   "Carrier_60_G120DStatusWord.12" AT %I3363.4 : Bool;   // Bit_12_BRAKE_OPEN
   "Carrier_60_G120DStatusWord.13" AT %I3363.5 : Bool;   // Bit_13_NO_OVERTEMP
   "Carrier_60_G120DStatusWord.14" AT %I3363.6 : Bool;   // Bit_14_CW_CCW
   "Carrier_60_G120DStatusWord.15" AT %I3363.7 : Bool;   // Bit_15_OVERL
   "Carrier_60_Slot2_Input" AT %IW3364 : Word;   // SLOT 2 INPUT WORD
   "Carrier_60_CrashDetectSW" AT %I3364.0 : Bool;   // CRASH DETECT SW
   "Carrier_60_SpareSafetyInput(2_1)" AT %I3364.1 : Bool;   // SPARE SAFETY INPUT
   "Carrier_60_SpareSafetyInput(2_2)" AT %I3364.2 : Bool;   // SPARE SAFETY INPUT
   "Carrier_60_SpareSafetyInput(2_3)" AT %I3364.3 : Bool;   // SPARE SAFETY INPUT
   "Carrier_60_SpareSafetyInput(2_4)" AT %I3364.4 : Bool;   // SPARE SAFETY INPUT
   "Carrier_60_SpareSafetyInput(2_5)" AT %I3364.5 : Bool;   // SPARE SAFETY INPUT
   "Carrier_60_SpareSafetyInput(2_6)" AT %I3364.6 : Bool;   // SPARE SAFETY INPUT
   "Carrier_60_SpareSafetyInput(2_7)" AT %I3364.7 : Bool;   // SPARE SAFETY INPUT
   "Carrier_60_Slot3_SafetyOutput" AT %IW3365 : Word;   // SLOT 3 SAFETY OUTPUT WORD
   "Carrier_60_Crash_Detect_OK" AT %I3365.0 : Bool;   // CARRIER CRASH DETECT
   "Carrier_60_SpareSafetyOutput(3_1)" AT %I3365.1 : Bool;   // SPARE SAFETY OUTPUT
   "Carrier_60_SpareSafetyOutput(3_2)" AT %I3365.2 : Bool;   // SPARE SAFETY OUTPUT
   "Carrier_60_SpareSafetyOutput(3_3)" AT %I3365.3 : Bool;   // SPARE SAFETY OUTPUT
   "Carrier_60_SpareSafetyOutput(3_4)" AT %I3365.4 : Bool;   // SPARE SAFETY OUTPUT
   "Carrier_60_SpareSafetyOutput(3_5)" AT %I3365.5 : Bool;   // SPARE SAFETY OUTPUT
   "Carrier_60_SpareSafetyOutput(3_6)" AT %I3365.6 : Bool;   // SPARE SAFETY OUTPUT
   "Carrier_60_SpareSafetyOutput(3_7)" AT %I3365.7 : Bool;   // SPARE SAFETY OUTPUT
   "Carrier_60_Slot4_Input" AT %IW3366 : Word;   // SLOT 4 INPUT WORD
   "Carrier_60_480VPowerOn_MDCB1" AT %I3366.0 : Bool;   // 480 VAC POWER ON MDCB 1
   "Carrier_60_SpareInput(4_1)" AT %I3366.1 : Bool;   // SPARE INPUT
   "Carrier_60_SpareInput(4_2)" AT %I3366.2 : Bool;   // SPARE INPUT
   "Carrier_60_SitopSelectStatus" AT %I3366.3 : Bool;   // SITOP SELECT STATUS
   "Carrier_60_DCsupplyOnPSCB2" AT %I3366.4 : Bool;   // DC SUPPLY ON PSCB 2
   "Carrier_60_SpareInput(4_5)" AT %I3366.5 : Bool;   // SPARE INPUT
   "Carrier_60_SpareInput(4_6)" AT %I3366.6 : Bool;   // SPARE INPUT
   "Carrier_60_SpareInput(4_7)" AT %I3366.7 : Bool;   // SPARE INPUT
   "Carrier_60_PB1_ProdHoldLH" AT %I3367.0 : Bool;   // PB 1 PRODUCTION HOLD LH
   "Carrier_60_PB2_ResetLH" AT %I3367.1 : Bool;   // PB 2 RESET LH
   "Carrier_60_PB3_ProdHoldRH" AT %I3367.2 : Bool;   // PB 3 PRODUCTION HOLD RH
   "Carrier_60_PB4_ResetRH" AT %I3367.3 : Bool;   // PB 4 RESET RH
   "Carrier_60_SpareInput(4_14)" AT %I3367.4 : Bool;   // SPARE INPUT
   "Carrier_60_SpareInput(4_15)" AT %I3367.5 : Bool;   // SPARE INPUT
   "Carrier_60_SpareInput(4_16)" AT %I3367.6 : Bool;   // SPARE INPUT
   "Carrier_60_SpareInput(4_17)" AT %I3367.7 : Bool;   // SPARE INPUT
   "Carrier_60_Slot5_Output" AT %IW3368 : Word;   // SLOT 5 OUTPUT WORD
   "Carrier_60_IRD400_HMI_24VDC_ENABLE" AT %I3368.0 : Bool;   // IRD 400 PANEL HMI 24V DC POWER
   "Carrier_60_FaultLight_LH" AT %I3368.1 : Bool;   // FAULT LIGHT LH
   "Carrier_60_RunLight_LH" AT %I3368.2 : Bool;   // RUN LIGHT LH
   "Carrier_60_FaultLight_RH" AT %I3368.3 : Bool;   // FAULT LIGHT RH
   "Carrier_60_RunLight_RH" AT %I3368.4 : Bool;   // RUN LIGHT RH
   "Carrier_60_SpareOutput(5_5)" AT %I3368.5 : Bool;   // SPARE OUTPUT
   "Carrier_60_SpareOutput(5_6)" AT %I3368.6 : Bool;   // SPARE OUTPUT
   "Carrier_60_SpareOutput(5_7)" AT %I3368.7 : Bool;   // SPARE OUTPUT
   "Carrier_60_ActualSpeed" AT %IW3370 : Word;   // ACTUAL SPEED
   "Carrier_60_CarrierDriveAlarm" AT %IW3372 : Word;   // CARRIER DRIVE ALARM
   "Carrier_60_CarrierDriveWarning" AT %IW3374 : Word;   // CARRIER DRIVE WARNING
   "Carrier_61_Status" AT %IW3400 : Word;   // CARRIER STATUS WORD
   "Carrier_61_Status.0" AT %I3400.0 : Bool;   // HEARTBEAT
   "Carrier_61_Status.1" AT %I3400.1 : Bool;   // MANUAL
   "Carrier_61_Status.2" AT %I3400.2 : Bool;   // IN_AUTO
   "Carrier_61_Status.3" AT %I3400.3 : Bool;   // POSITIONING_COMPLETE
   "Carrier_61_Status.4" AT %I3400.4 : Bool;   // PRODUCTION HOLD
   "Carrier_61_Status.5" AT %I3400.5 : Bool;   // CARRIER MOVING FORWARD
   "Carrier_61_Status.6" AT %I3400.6 : Bool;   // CARRIER MOVING REVERSE
   "Carrier_61_Status.7" AT %I3400.7 : Bool;   // CARRIER FAULT
   "Carrier_61_Status.8" AT %I3401.0 : Bool;   // CRASH DETECT TRIPPED
   "Carrier_61_Status.9" AT %I3401.1 : Bool;
   "Carrier_61_Status.10" AT %I3401.2 : Bool;
   "Carrier_61_Status.11" AT %I3401.3 : Bool;
   "Carrier_61_Status.12" AT %I3401.4 : Bool;
   "Carrier_61_Status.13" AT %I3401.5 : Bool;
   "Carrier_61_Status.14" AT %I3401.6 : Bool;
   "Carrier_61_Status.15" AT %I3401.7 : Bool;
   "Carrier_61_SDCFaultCode" AT %IW3402 : Word;   // SDC FAULT CODE
   "Carrier_61_CarrierPosition" AT %ID3404 : DWord;   // CARRIER POSITION
   "Carrier_61_CarrierNumber" AT %IW3408 : Word;   // CARRIER NUMBER
   "Carrier_61_G120DControlWord" AT %IW3410 : Word;   // G120D_STW1_CONTROL
   "Carrier_61_G120DControlWord.0" AT %I3410.0 : Bool;   // Bit_00_ON
   "Carrier_61_G120DControlWord.1" AT %I3410.1 : Bool;   // Bit_01_AUS2_INH
   "Carrier_61_G120DControlWord.2" AT %I3410.2 : Bool;   // Bit_02_AUS3_STOP
   "Carrier_61_G120DControlWord.3" AT %I3410.3 : Bool;   // Bit_03_EN
   "Carrier_61_G120DControlWord.4" AT %I3410.4 : Bool;   // Bit_04_EN_RAMP
   "Carrier_61_G120DControlWord.5" AT %I3410.5 : Bool;   // Bit_05_START_RAMP
   "Carrier_61_G120DControlWord.6" AT %I3410.6 : Bool;   // Bit_06_SETPOINT
   "Carrier_61_G120DControlWord.7" AT %I3410.7 : Bool;   // Bit_07_RESET
   "Carrier_61_G120DControlWord.8" AT %I3411.0 : Bool;   // Bit_08_JOG_R
   "Carrier_61_G120DControlWord.9" AT %I3411.1 : Bool;   // Bit_09_JOG_L
   "Carrier_61_G120DControlWord.10" AT %I3411.2 : Bool;   // Bit_10_CONTR_PLC
   "Carrier_61_G120DControlWord.11" AT %I3411.3 : Bool;   // Bit_11_REVERSE
   "Carrier_61_G120DControlWord.12" AT %I3411.4 : Bool;   // Bit_12_BRAKE_RELEASE
   "Carrier_61_G120DControlWord.13" AT %I3411.5 : Bool;   // Bit_13_DDS
   "Carrier_61_G120DControlWord.14" AT %I3411.6 : Bool;   // Bit_14_DO0
   "Carrier_61_G120DControlWord.15" AT %I3411.7 : Bool;   // Bit_15_DO1
   "Carrier_61_G120DStatusWord" AT %IW3412 : Word;   // G120D_ZSW1_STATUS
   "Carrier_61_G120DStatusWord.0" AT %I3412.0 : Bool;   // Bit_00_READY_RUN
   "Carrier_61_G120DStatusWord.1" AT %I3412.1 : Bool;   // Bit_01_READY_ON
   "Carrier_61_G120DStatusWord.2" AT %I3412.2 : Bool;   // Bit_02_ENABLE
   "Carrier_61_G120DStatusWord.3" AT %I3412.3 : Bool;   // Bit_03_FAULT
   "Carrier_61_G120DStatusWord.4" AT %I3412.4 : Bool;   // Bit_04_OFF2
   "Carrier_61_G120DStatusWord.5" AT %I3412.5 : Bool;   // Bit_05_OFF3
   "Carrier_61_G120DStatusWord.6" AT %I3412.6 : Bool;   // Bit_06_LOCK_OUT
   "Carrier_61_G120DStatusWord.7" AT %I3412.7 : Bool;   // Bit_07_WARN
   "Carrier_61_G120DStatusWord.8" AT %I3413.0 : Bool;   // Bit_08_NO_DEVIATION
   "Carrier_61_G120DStatusWord.9" AT %I3413.1 : Bool;   // Bit_09_CONTR_PLC
   "Carrier_61_G120DStatusWord.10" AT %I3413.2 : Bool;   // Bit_10_F_MAX
   "Carrier_61_G120DStatusWord.11" AT %I3413.3 : Bool;   // Bit_11_LIMIT_REACHED
   "Carrier_61_G120DStatusWord.12" AT %I3413.4 : Bool;   // Bit_12_BRAKE_OPEN
   "Carrier_61_G120DStatusWord.13" AT %I3413.5 : Bool;   // Bit_13_NO_OVERTEMP
   "Carrier_61_G120DStatusWord.14" AT %I3413.6 : Bool;   // Bit_14_CW_CCW
   "Carrier_61_G120DStatusWord.15" AT %I3413.7 : Bool;   // Bit_15_OVERL
   "Carrier_61_Slot2_Input" AT %IW3414 : Word;   // SLOT 2 INPUT WORD
   "Carrier_61_CrashDetectSW" AT %I3414.0 : Bool;   // CRASH DETECT SW
   "Carrier_61_SpareSafetyInput(2_1)" AT %I3414.1 : Bool;   // SPARE SAFETY INPUT
   "Carrier_61_SpareSafetyInput(2_2)" AT %I3414.2 : Bool;   // SPARE SAFETY INPUT
   "Carrier_61_SpareSafetyInput(2_3)" AT %I3414.3 : Bool;   // SPARE SAFETY INPUT
   "Carrier_61_SpareSafetyInput(2_4)" AT %I3414.4 : Bool;   // SPARE SAFETY INPUT
   "Carrier_61_SpareSafetyInput(2_5)" AT %I3414.5 : Bool;   // SPARE SAFETY INPUT
   "Carrier_61_SpareSafetyInput(2_6)" AT %I3414.6 : Bool;   // SPARE SAFETY INPUT
   "Carrier_61_SpareSafetyInput(2_7)" AT %I3414.7 : Bool;   // SPARE SAFETY INPUT
   "Carrier_61_Slot3_SafetyOutput" AT %IW3415 : Word;   // SLOT 3 SAFETY OUTPUT WORD
   "Carrier_61_Crash_Detect_OK" AT %I3415.0 : Bool;   // CARRIER CRASH DETECT
   "Carrier_61_SpareSafetyOutput(3_1)" AT %I3415.1 : Bool;   // SPARE SAFETY OUTPUT
   "Carrier_61_SpareSafetyOutput(3_2)" AT %I3415.2 : Bool;   // SPARE SAFETY OUTPUT
   "Carrier_61_SpareSafetyOutput(3_3)" AT %I3415.3 : Bool;   // SPARE SAFETY OUTPUT
   "Carrier_61_SpareSafetyOutput(3_4)" AT %I3415.4 : Bool;   // SPARE SAFETY OUTPUT
   "Carrier_61_SpareSafetyOutput(3_5)" AT %I3415.5 : Bool;   // SPARE SAFETY OUTPUT
   "Carrier_61_SpareSafetyOutput(3_6)" AT %I3415.6 : Bool;   // SPARE SAFETY OUTPUT
   "Carrier_61_SpareSafetyOutput(3_7)" AT %I3415.7 : Bool;   // SPARE SAFETY OUTPUT
   "Carrier_61_Slot4_Input" AT %IW3416 : Word;   // SLOT 4 INPUT WORD
   "Carrier_61_480VPowerOn_MDCB1" AT %I3416.0 : Bool;   // 480 VAC POWER ON MDCB 1
   "Carrier_61_SpareInput(4_1)" AT %I3416.1 : Bool;   // SPARE INPUT
   "Carrier_61_SpareInput(4_2)" AT %I3416.2 : Bool;   // SPARE INPUT
   "Carrier_61_SitopSelectStatus" AT %I3416.3 : Bool;   // SITOP SELECT STATUS
   "Carrier_61_DCsupplyOnPSCB2" AT %I3416.4 : Bool;   // DC SUPPLY ON PSCB 2
   "Carrier_61_SpareInput(4_5)" AT %I3416.5 : Bool;   // SPARE INPUT
   "Carrier_61_SpareInput(4_6)" AT %I3416.6 : Bool;   // SPARE INPUT
   "Carrier_61_SpareInput(4_7)" AT %I3416.7 : Bool;   // SPARE INPUT
   "Carrier_61_PB1_ProdHoldLH" AT %I3417.0 : Bool;   // PB 1 PRODUCTION HOLD LH
   "Carrier_61_PB2_ResetLH" AT %I3417.1 : Bool;   // PB 2 RESET LH
   "Carrier_61_PB3_ProdHoldRH" AT %I3417.2 : Bool;   // PB 3 PRODUCTION HOLD RH
   "Carrier_61_PB4_ResetRH" AT %I3417.3 : Bool;   // PB 4 RESET RH
   "Carrier_61_SpareInput(4_14)" AT %I3417.4 : Bool;   // SPARE INPUT
   "Carrier_61_SpareInput(4_15)" AT %I3417.5 : Bool;   // SPARE INPUT
   "Carrier_61_SpareInput(4_16)" AT %I3417.6 : Bool;   // SPARE INPUT
   "Carrier_61_SpareInput(4_17)" AT %I3417.7 : Bool;   // SPARE INPUT
   "Carrier_61_Slot5_Output" AT %IW3418 : Word;   // SLOT 5 OUTPUT WORD
   "Carrier_61_IRD400_HMI_24VDC_ENABLE" AT %I3418.0 : Bool;   // IRD 400 PANEL HMI 24V DC POWER
   "Carrier_61_FaultLight_LH" AT %I3418.1 : Bool;   // FAULT LIGHT LH
   "Carrier_61_RunLight_LH" AT %I3418.2 : Bool;   // RUN LIGHT LH
   "Carrier_61_FaultLight_RH" AT %I3418.3 : Bool;   // FAULT LIGHT RH
   "Carrier_61_RunLight_RH" AT %I3418.4 : Bool;   // RUN LIGHT RH
   "Carrier_61_SpareOutput(5_5)" AT %I3418.5 : Bool;   // SPARE OUTPUT
   "Carrier_61_SpareOutput(5_6)" AT %I3418.6 : Bool;   // SPARE OUTPUT
   "Carrier_61_SpareOutput(5_7)" AT %I3418.7 : Bool;   // SPARE OUTPUT
   "Carrier_61_ActualSpeed" AT %IW3420 : Word;   // ACTUAL SPEED
   "Carrier_61_CarrierDriveAlarm" AT %IW3422 : Word;   // CARRIER DRIVE ALARM
   "Carrier_61_CarrierDriveWarning" AT %IW3424 : Word;   // CARRIER DRIVE WARNING
   "Carrier_62_Status" AT %IW3450 : Word;   // CARRIER STATUS WORD
   "Carrier_62_Status.0" AT %I3450.0 : Bool;   // HEARTBEAT
   "Carrier_62_Status.1" AT %I3450.1 : Bool;   // MANUAL
   "Carrier_62_Status.2" AT %I3450.2 : Bool;   // IN_AUTO
   "Carrier_62_Status.3" AT %I3450.3 : Bool;   // POSITIONING_COMPLETE
   "Carrier_62_Status.4" AT %I3450.4 : Bool;   // PRODUCTION HOLD
   "Carrier_62_Status.5" AT %I3450.5 : Bool;   // CARRIER MOVING FORWARD
   "Carrier_62_Status.6" AT %I3450.6 : Bool;   // CARRIER MOVING REVERSE
   "Carrier_62_Status.7" AT %I3450.7 : Bool;   // CARRIER FAULT
   "Carrier_62_Status.8" AT %I3451.0 : Bool;   // CRASH DETECT TRIPPED
   "Carrier_62_Status.9" AT %I3451.1 : Bool;
   "Carrier_62_Status.10" AT %I3451.2 : Bool;
   "Carrier_62_Status.11" AT %I3451.3 : Bool;
   "Carrier_62_Status.12" AT %I3451.4 : Bool;
   "Carrier_62_Status.13" AT %I3451.5 : Bool;
   "Carrier_62_Status.14" AT %I3451.6 : Bool;
   "Carrier_62_Status.15" AT %I3451.7 : Bool;
   "Carrier_62_SDCFaultCode" AT %IW3452 : Word;   // SDC FAULT CODE
   "Carrier_62_CarrierPosition" AT %ID3454 : DWord;   // CARRIER POSITION
   "Carrier_62_CarrierNumber" AT %IW3458 : Word;   // CARRIER NUMBER
   "Carrier_62_G120DControlWord" AT %IW3460 : Word;   // G120D_STW1_CONTROL
   "Carrier_62_G120DControlWord.0" AT %I3460.0 : Bool;   // Bit_00_ON
   "Carrier_62_G120DControlWord.1" AT %I3460.1 : Bool;   // Bit_01_AUS2_INH
   "Carrier_62_G120DControlWord.2" AT %I3460.2 : Bool;   // Bit_02_AUS3_STOP
   "Carrier_62_G120DControlWord.3" AT %I3460.3 : Bool;   // Bit_03_EN
   "Carrier_62_G120DControlWord.4" AT %I3460.4 : Bool;   // Bit_04_EN_RAMP
   "Carrier_62_G120DControlWord.5" AT %I3460.5 : Bool;   // Bit_05_START_RAMP
   "Carrier_62_G120DControlWord.6" AT %I3460.6 : Bool;   // Bit_06_SETPOINT
   "Carrier_62_G120DControlWord.7" AT %I3460.7 : Bool;   // Bit_07_RESET
   "Carrier_62_G120DControlWord.8" AT %I3461.0 : Bool;   // Bit_08_JOG_R
   "Carrier_62_G120DControlWord.9" AT %I3461.1 : Bool;   // Bit_09_JOG_L
   "Carrier_62_G120DControlWord.10" AT %I3461.2 : Bool;   // Bit_10_CONTR_PLC
   "Carrier_62_G120DControlWord.11" AT %I3461.3 : Bool;   // Bit_11_REVERSE
   "Carrier_62_G120DControlWord.12" AT %I3461.4 : Bool;   // Bit_12_BRAKE_RELEASE
   "Carrier_62_G120DControlWord.13" AT %I3461.5 : Bool;   // Bit_13_DDS
   "Carrier_62_G120DControlWord.14" AT %I3461.6 : Bool;   // Bit_14_DO0
   "Carrier_62_G120DControlWord.15" AT %I3461.7 : Bool;   // Bit_15_DO1
   "Carrier_62_G120DStatusWord" AT %IW3462 : Word;   // G120D_ZSW1_STATUS
   "Carrier_62_G120DStatusWord.0" AT %I3462.0 : Bool;   // Bit_00_READY_RUN
   "Carrier_62_G120DStatusWord.1" AT %I3462.1 : Bool;   // Bit_01_READY_ON
   "Carrier_62_G120DStatusWord.2" AT %I3462.2 : Bool;   // Bit_02_ENABLE
   "Carrier_62_G120DStatusWord.3" AT %I3462.3 : Bool;   // Bit_03_FAULT
   "Carrier_62_G120DStatusWord.4" AT %I3462.4 : Bool;   // Bit_04_OFF2
   "Carrier_62_G120DStatusWord.5" AT %I3462.5 : Bool;   // Bit_05_OFF3
   "Carrier_62_G120DStatusWord.6" AT %I3462.6 : Bool;   // Bit_06_LOCK_OUT
   "Carrier_62_G120DStatusWord.7" AT %I3462.7 : Bool;   // Bit_07_WARN
   "Carrier_62_G120DStatusWord.8" AT %I3463.0 : Bool;   // Bit_08_NO_DEVIATION
   "Carrier_62_G120DStatusWord.9" AT %I3463.1 : Bool;   // Bit_09_CONTR_PLC
   "Carrier_62_G120DStatusWord.10" AT %I3463.2 : Bool;   // Bit_10_F_MAX
   "Carrier_62_G120DStatusWord.11" AT %I3463.3 : Bool;   // Bit_11_LIMIT_REACHED
   "Carrier_62_G120DStatusWord.12" AT %I3463.4 : Bool;   // Bit_12_BRAKE_OPEN
   "Carrier_62_G120DStatusWord.13" AT %I3463.5 : Bool;   // Bit_13_NO_OVERTEMP
   "Carrier_62_G120DStatusWord.14" AT %I3463.6 : Bool;   // Bit_14_CW_CCW
   "Carrier_62_G120DStatusWord.15" AT %I3463.7 : Bool;   // Bit_15_OVERL
   "Carrier_62_Slot2_Input" AT %IW3464 : Word;   // SLOT 2 INPUT WORD
   "Carrier_62_CrashDetectSW" AT %I3464.0 : Bool;   // CRASH DETECT SW
   "Carrier_62_SpareSafetyInput(2_1)" AT %I3464.1 : Bool;   // SPARE SAFETY INPUT
   "Carrier_62_SpareSafetyInput(2_2)" AT %I3464.2 : Bool;   // SPARE SAFETY INPUT
   "Carrier_62_SpareSafetyInput(2_3)" AT %I3464.3 : Bool;   // SPARE SAFETY INPUT
   "Carrier_62_SpareSafetyInput(2_4)" AT %I3464.4 : Bool;   // SPARE SAFETY INPUT
   "Carrier_62_SpareSafetyInput(2_5)" AT %I3464.5 : Bool;   // SPARE SAFETY INPUT
   "Carrier_62_SpareSafetyInput(2_6)" AT %I3464.6 : Bool;   // SPARE SAFETY INPUT
   "Carrier_62_SpareSafetyInput(2_7)" AT %I3464.7 : Bool;   // SPARE SAFETY INPUT
   "Carrier_62_Slot3_SafetyOutput" AT %IW3465 : Word;   // SLOT 3 SAFETY OUTPUT WORD
   "Carrier_62_Crash_Detect_OK" AT %I3465.0 : Bool;   // CARRIER CRASH DETECT
   "Carrier_62_SpareSafetyOutput(3_1)" AT %I3465.1 : Bool;   // SPARE SAFETY OUTPUT
   "Carrier_62_SpareSafetyOutput(3_2)" AT %I3465.2 : Bool;   // SPARE SAFETY OUTPUT
   "Carrier_62_SpareSafetyOutput(3_3)" AT %I3465.3 : Bool;   // SPARE SAFETY OUTPUT
   "Carrier_62_SpareSafetyOutput(3_4)" AT %I3465.4 : Bool;   // SPARE SAFETY OUTPUT
   "Carrier_62_SpareSafetyOutput(3_5)" AT %I3465.5 : Bool;   // SPARE SAFETY OUTPUT
   "Carrier_62_SpareSafetyOutput(3_6)" AT %I3465.6 : Bool;   // SPARE SAFETY OUTPUT
   "Carrier_62_SpareSafetyOutput(3_7)" AT %I3465.7 : Bool;   // SPARE SAFETY OUTPUT
   "Carrier_62_Slot4_Input" AT %IW3466 : Word;   // SLOT 4 INPUT WORD
   "Carrier_62_480VPowerOn_MDCB1" AT %I3466.0 : Bool;   // 480 VAC POWER ON MDCB 1
   "Carrier_62_SpareInput(4_1)" AT %I3466.1 : Bool;   // SPARE INPUT
   "Carrier_62_SpareInput(4_2)" AT %I3466.2 : Bool;   // SPARE INPUT
   "Carrier_62_SitopSelectStatus" AT %I3466.3 : Bool;   // SITOP SELECT STATUS
   "Carrier_62_DCsupplyOnPSCB2" AT %I3466.4 : Bool;   // DC SUPPLY ON PSCB 2
   "Carrier_62_SpareInput(4_5)" AT %I3466.5 : Bool;   // SPARE INPUT
   "Carrier_62_SpareInput(4_6)" AT %I3466.6 : Bool;   // SPARE INPUT
   "Carrier_62_SpareInput(4_7)" AT %I3466.7 : Bool;   // SPARE INPUT
   "Carrier_62_PB1_ProdHoldLH" AT %I3467.0 : Bool;   // PB 1 PRODUCTION HOLD LH
   "Carrier_62_PB2_ResetLH" AT %I3467.1 : Bool;   // PB 2 RESET LH
   "Carrier_62_PB3_ProdHoldRH" AT %I3467.2 : Bool;   // PB 3 PRODUCTION HOLD RH
   "Carrier_62_PB4_ResetRH" AT %I3467.3 : Bool;   // PB 4 RESET RH
   "Carrier_62_SpareInput(4_14)" AT %I3467.4 : Bool;   // SPARE INPUT
   "Carrier_62_SpareInput(4_15)" AT %I3467.5 : Bool;   // SPARE INPUT
   "Carrier_62_SpareInput(4_16)" AT %I3467.6 : Bool;   // SPARE INPUT
   "Carrier_62_SpareInput(4_17)" AT %I3467.7 : Bool;   // SPARE INPUT
   "Carrier_62_Slot5_Output" AT %IW3468 : Word;   // SLOT 5 OUTPUT WORD
   "Carrier_62_IRD400_HMI_24VDC_ENABLE" AT %I3468.0 : Bool;   // IRD 400 PANEL HMI 24V DC POWER
   "Carrier_62_FaultLight_LH" AT %I3468.1 : Bool;   // FAULT LIGHT LH
   "Carrier_62_RunLight_LH" AT %I3468.2 : Bool;   // RUN LIGHT LH
   "Carrier_62_FaultLight_RH" AT %I3468.3 : Bool;   // FAULT LIGHT RH
   "Carrier_62_RunLight_RH" AT %I3468.4 : Bool;   // RUN LIGHT RH
   "Carrier_62_SpareOutput(5_5)" AT %I3468.5 : Bool;   // SPARE OUTPUT
   "Carrier_62_SpareOutput(5_6)" AT %I3468.6 : Bool;   // SPARE OUTPUT
   "Carrier_62_SpareOutput(5_7)" AT %I3468.7 : Bool;   // SPARE OUTPUT
   "Carrier_62_ActualSpeed" AT %IW3470 : Word;   // ACTUAL SPEED
   "Carrier_62_CarrierDriveAlarm" AT %IW3472 : Word;   // CARRIER DRIVE ALARM
   "Carrier_62_CarrierDriveWarning" AT %IW3474 : Word;   // CARRIER DRIVE WARNING
   "Carrier_63_Status" AT %IW3500 : Word;   // CARRIER STATUS WORD
   "Carrier_63_Status.0" AT %I3500.0 : Bool;   // HEARTBEAT
   "Carrier_63_Status.1" AT %I3500.1 : Bool;   // MANUAL
   "Carrier_63_Status.2" AT %I3500.2 : Bool;   // IN_AUTO
   "Carrier_63_Status.3" AT %I3500.3 : Bool;   // POSITIONING_COMPLETE
   "Carrier_63_Status.4" AT %I3500.4 : Bool;   // PRODUCTION HOLD
   "Carrier_63_Status.5" AT %I3500.5 : Bool;   // CARRIER MOVING FORWARD
   "Carrier_63_Status.6" AT %I3500.6 : Bool;   // CARRIER MOVING REVERSE
   "Carrier_63_Status.7" AT %I3500.7 : Bool;   // CARRIER FAULT
   "Carrier_63_Status.8" AT %I3501.0 : Bool;   // CRASH DETECT TRIPPED
   "Carrier_63_Status.9" AT %I3501.1 : Bool;
   "Carrier_63_Status.10" AT %I3501.2 : Bool;
   "Carrier_63_Status.11" AT %I3501.3 : Bool;
   "Carrier_63_Status.12" AT %I3501.4 : Bool;
   "Carrier_63_Status.13" AT %I3501.5 : Bool;
   "Carrier_63_Status.14" AT %I3501.6 : Bool;
   "Carrier_63_Status.15" AT %I3501.7 : Bool;
   "Carrier_63_SDCFaultCode" AT %IW3502 : Word;   // SDC FAULT CODE
   "Carrier_63_CarrierPosition" AT %ID3504 : DWord;   // CARRIER POSITION
   "Carrier_63_CarrierNumber" AT %IW3508 : Word;   // CARRIER NUMBER
   "Carrier_63_G120DControlWord" AT %IW3510 : Word;   // G120D_STW1_CONTROL
   "Carrier_63_G120DControlWord.0" AT %I3510.0 : Bool;   // Bit_00_ON
   "Carrier_63_G120DControlWord.1" AT %I3510.1 : Bool;   // Bit_01_AUS2_INH
   "Carrier_63_G120DControlWord.2" AT %I3510.2 : Bool;   // Bit_02_AUS3_STOP
   "Carrier_63_G120DControlWord.3" AT %I3510.3 : Bool;   // Bit_03_EN
   "Carrier_63_G120DControlWord.4" AT %I3510.4 : Bool;   // Bit_04_EN_RAMP
   "Carrier_63_G120DControlWord.5" AT %I3510.5 : Bool;   // Bit_05_START_RAMP
   "Carrier_63_G120DControlWord.6" AT %I3510.6 : Bool;   // Bit_06_SETPOINT
   "Carrier_63_G120DControlWord.7" AT %I3510.7 : Bool;   // Bit_07_RESET
   "Carrier_63_G120DControlWord.8" AT %I3511.0 : Bool;   // Bit_08_JOG_R
   "Carrier_63_G120DControlWord.9" AT %I3511.1 : Bool;   // Bit_09_JOG_L
   "Carrier_63_G120DControlWord.10" AT %I3511.2 : Bool;   // Bit_10_CONTR_PLC
   "Carrier_63_G120DControlWord.11" AT %I3511.3 : Bool;   // Bit_11_REVERSE
   "Carrier_63_G120DControlWord.12" AT %I3511.4 : Bool;   // Bit_12_BRAKE_RELEASE
   "Carrier_63_G120DControlWord.13" AT %I3511.5 : Bool;   // Bit_13_DDS
   "Carrier_63_G120DControlWord.14" AT %I3511.6 : Bool;   // Bit_14_DO0
   "Carrier_63_G120DControlWord.15" AT %I3511.7 : Bool;   // Bit_15_DO1
   "Carrier_63_G120DStatusWord" AT %IW3512 : Word;   // G120D_ZSW1_STATUS
   "Carrier_63_G120DStatusWord.0" AT %I3512.0 : Bool;   // Bit_00_READY_RUN
   "Carrier_63_G120DStatusWord.1" AT %I3512.1 : Bool;   // Bit_01_READY_ON
   "Carrier_63_G120DStatusWord.2" AT %I3512.2 : Bool;   // Bit_02_ENABLE
   "Carrier_63_G120DStatusWord.3" AT %I3512.3 : Bool;   // Bit_03_FAULT
   "Carrier_63_G120DStatusWord.4" AT %I3512.4 : Bool;   // Bit_04_OFF2
   "Carrier_63_G120DStatusWord.5" AT %I3512.5 : Bool;   // Bit_05_OFF3
   "Carrier_63_G120DStatusWord.6" AT %I3512.6 : Bool;   // Bit_06_LOCK_OUT
   "Carrier_63_G120DStatusWord.7" AT %I3512.7 : Bool;   // Bit_07_WARN
   "Carrier_63_G120DStatusWord.8" AT %I3513.0 : Bool;   // Bit_08_NO_DEVIATION
   "Carrier_63_G120DStatusWord.9" AT %I3513.1 : Bool;   // Bit_09_CONTR_PLC
   "Carrier_63_G120DStatusWord.10" AT %I3513.2 : Bool;   // Bit_10_F_MAX
   "Carrier_63_G120DStatusWord.11" AT %I3513.3 : Bool;   // Bit_11_LIMIT_REACHED
   "Carrier_63_G120DStatusWord.12" AT %I3513.4 : Bool;   // Bit_12_BRAKE_OPEN
   "Carrier_63_G120DStatusWord.13" AT %I3513.5 : Bool;   // Bit_13_NO_OVERTEMP
   "Carrier_63_G120DStatusWord.14" AT %I3513.6 : Bool;   // Bit_14_CW_CCW
   "Carrier_63_G120DStatusWord.15" AT %I3513.7 : Bool;   // Bit_15_OVERL
   "Carrier_63_Slot2_Input" AT %IW3514 : Word;   // SLOT 2 INPUT WORD
   "Carrier_63_CrashDetectSW" AT %I3514.0 : Bool;   // CRASH DETECT SW
   "Carrier_63_SpareSafetyInput(2_1)" AT %I3514.1 : Bool;   // SPARE SAFETY INPUT
   "Carrier_63_SpareSafetyInput(2_2)" AT %I3514.2 : Bool;   // SPARE SAFETY INPUT
   "Carrier_63_SpareSafetyInput(2_3)" AT %I3514.3 : Bool;   // SPARE SAFETY INPUT
   "Carrier_63_SpareSafetyInput(2_4)" AT %I3514.4 : Bool;   // SPARE SAFETY INPUT
   "Carrier_63_SpareSafetyInput(2_5)" AT %I3514.5 : Bool;   // SPARE SAFETY INPUT
   "Carrier_63_SpareSafetyInput(2_6)" AT %I3514.6 : Bool;   // SPARE SAFETY INPUT
   "Carrier_63_SpareSafetyInput(2_7)" AT %I3514.7 : Bool;   // SPARE SAFETY INPUT
   "Carrier_63_Slot3_SafetyOutput" AT %IW3515 : Word;   // SLOT 3 SAFETY OUTPUT WORD
   "Carrier_63_Crash_Detect_OK" AT %I3515.0 : Bool;   // CARRIER CRASH DETECT
   "Carrier_63_SpareSafetyOutput(3_1)" AT %I3515.1 : Bool;   // SPARE SAFETY OUTPUT
   "Carrier_63_SpareSafetyOutput(3_2)" AT %I3515.2 : Bool;   // SPARE SAFETY OUTPUT
   "Carrier_63_SpareSafetyOutput(3_3)" AT %I3515.3 : Bool;   // SPARE SAFETY OUTPUT
   "Carrier_63_SpareSafetyOutput(3_4)" AT %I3515.4 : Bool;   // SPARE SAFETY OUTPUT
   "Carrier_63_SpareSafetyOutput(3_5)" AT %I3515.5 : Bool;   // SPARE SAFETY OUTPUT
   "Carrier_63_SpareSafetyOutput(3_6)" AT %I3515.6 : Bool;   // SPARE SAFETY OUTPUT
   "Carrier_63_SpareSafetyOutput(3_7)" AT %I3515.7 : Bool;   // SPARE SAFETY OUTPUT
   "Carrier_63_Slot4_Input" AT %IW3516 : Word;   // SLOT 4 INPUT WORD
   "Carrier_63_480VPowerOn_MDCB1" AT %I3516.0 : Bool;   // 480 VAC POWER ON MDCB 1
   "Carrier_63_SpareInput(4_1)" AT %I3516.1 : Bool;   // SPARE INPUT
   "Carrier_63_SpareInput(4_2)" AT %I3516.2 : Bool;   // SPARE INPUT
   "Carrier_63_SitopSelectStatus" AT %I3516.3 : Bool;   // SITOP SELECT STATUS
   "Carrier_63_DCsupplyOnPSCB2" AT %I3516.4 : Bool;   // DC SUPPLY ON PSCB 2
   "Carrier_63_SpareInput(4_5)" AT %I3516.5 : Bool;   // SPARE INPUT
   "Carrier_63_SpareInput(4_6)" AT %I3516.6 : Bool;   // SPARE INPUT
   "Carrier_63_SpareInput(4_7)" AT %I3516.7 : Bool;   // SPARE INPUT
   "Carrier_63_PB1_ProdHoldLH" AT %I3517.0 : Bool;   // PB 1 PRODUCTION HOLD LH
   "Carrier_63_PB2_ResetLH" AT %I3517.1 : Bool;   // PB 2 RESET LH
   "Carrier_63_PB3_ProdHoldRH" AT %I3517.2 : Bool;   // PB 3 PRODUCTION HOLD RH
   "Carrier_63_PB4_ResetRH" AT %I3517.3 : Bool;   // PB 4 RESET RH
   "Carrier_63_SpareInput(4_14)" AT %I3517.4 : Bool;   // SPARE INPUT
   "Carrier_63_SpareInput(4_15)" AT %I3517.5 : Bool;   // SPARE INPUT
   "Carrier_63_SpareInput(4_16)" AT %I3517.6 : Bool;   // SPARE INPUT
   "Carrier_63_SpareInput(4_17)" AT %I3517.7 : Bool;   // SPARE INPUT
   "Carrier_63_Slot5_Output" AT %IW3518 : Word;   // SLOT 5 OUTPUT WORD
   "Carrier_63_IRD400_HMI_24VDC_ENABLE" AT %I3518.0 : Bool;   // IRD 400 PANEL HMI 24V DC POWER
   "Carrier_63_FaultLight_LH" AT %I3518.1 : Bool;   // FAULT LIGHT LH
   "Carrier_63_RunLight_LH" AT %I3518.2 : Bool;   // RUN LIGHT LH
   "Carrier_63_FaultLight_RH" AT %I3518.3 : Bool;   // FAULT LIGHT RH
   "Carrier_63_RunLight_RH" AT %I3518.4 : Bool;   // RUN LIGHT RH
   "Carrier_63_SpareOutput(5_5)" AT %I3518.5 : Bool;   // SPARE OUTPUT
   "Carrier_63_SpareOutput(5_6)" AT %I3518.6 : Bool;   // SPARE OUTPUT
   "Carrier_63_SpareOutput(5_7)" AT %I3518.7 : Bool;   // SPARE OUTPUT
   "Carrier_63_ActualSpeed" AT %IW3520 : Word;   // ACTUAL SPEED
   "Carrier_63_CarrierDriveAlarm" AT %IW3522 : Word;   // CARRIER DRIVE ALARM
   "Carrier_63_CarrierDriveWarning" AT %IW3524 : Word;   // CARRIER DRIVE WARNING
   "Carrier_64_Status" AT %IW3550 : Word;   // CARRIER STATUS WORD
   "Carrier_64_Status.0" AT %I3550.0 : Bool;   // HEARTBEAT
   "Carrier_64_Status.1" AT %I3550.1 : Bool;   // MANUAL
   "Carrier_64_Status.2" AT %I3550.2 : Bool;   // IN_AUTO
   "Carrier_64_Status.3" AT %I3550.3 : Bool;   // POSITIONING_COMPLETE
   "Carrier_64_Status.4" AT %I3550.4 : Bool;   // PRODUCTION HOLD
   "Carrier_64_Status.5" AT %I3550.5 : Bool;   // CARRIER MOVING FORWARD
   "Carrier_64_Status.6" AT %I3550.6 : Bool;   // CARRIER MOVING REVERSE
   "Carrier_64_Status.7" AT %I3550.7 : Bool;   // CARRIER FAULT
   "Carrier_64_Status.8" AT %I3551.0 : Bool;   // CRASH DETECT TRIPPED
   "Carrier_64_Status.9" AT %I3551.1 : Bool;
   "Carrier_64_Status.10" AT %I3551.2 : Bool;
   "Carrier_64_Status.11" AT %I3551.3 : Bool;
   "Carrier_64_Status.12" AT %I3551.4 : Bool;
   "Carrier_64_Status.13" AT %I3551.5 : Bool;
   "Carrier_64_Status.14" AT %I3551.6 : Bool;
   "Carrier_64_Status.15" AT %I3551.7 : Bool;
   "Carrier_64_SDCFaultCode" AT %IW3552 : Word;   // SDC FAULT CODE
   "Carrier_64_CarrierPosition" AT %ID3554 : DWord;   // CARRIER POSITION
   "Carrier_64_CarrierNumber" AT %IW3558 : Word;   // CARRIER NUMBER
   "Carrier_64_G120DControlWord" AT %IW3560 : Word;   // G120D_STW1_CONTROL
   "Carrier_64_G120DControlWord.0" AT %I3560.0 : Bool;   // Bit_00_ON
   "Carrier_64_G120DControlWord.1" AT %I3560.1 : Bool;   // Bit_01_AUS2_INH
   "Carrier_64_G120DControlWord.2" AT %I3560.2 : Bool;   // Bit_02_AUS3_STOP
   "Carrier_64_G120DControlWord.3" AT %I3560.3 : Bool;   // Bit_03_EN
   "Carrier_64_G120DControlWord.4" AT %I3560.4 : Bool;   // Bit_04_EN_RAMP
   "Carrier_64_G120DControlWord.5" AT %I3560.5 : Bool;   // Bit_05_START_RAMP
   "Carrier_64_G120DControlWord.6" AT %I3560.6 : Bool;   // Bit_06_SETPOINT
   "Carrier_64_G120DControlWord.7" AT %I3560.7 : Bool;   // Bit_07_RESET
   "Carrier_64_G120DControlWord.8" AT %I3561.0 : Bool;   // Bit_08_JOG_R
   "Carrier_64_G120DControlWord.9" AT %I3561.1 : Bool;   // Bit_09_JOG_L
   "Carrier_64_G120DControlWord.10" AT %I3561.2 : Bool;   // Bit_10_CONTR_PLC
   "Carrier_64_G120DControlWord.11" AT %I3561.3 : Bool;   // Bit_11_REVERSE
   "Carrier_64_G120DControlWord.12" AT %I3561.4 : Bool;   // Bit_12_BRAKE_RELEASE
   "Carrier_64_G120DControlWord.13" AT %I3561.5 : Bool;   // Bit_13_DDS
   "Carrier_64_G120DControlWord.14" AT %I3561.6 : Bool;   // Bit_14_DO0
   "Carrier_64_G120DControlWord.15" AT %I3561.7 : Bool;   // Bit_15_DO1
   "Carrier_64_G120DStatusWord" AT %IW3562 : Word;   // G120D_ZSW1_STATUS
   "Carrier_64_G120DStatusWord.0" AT %I3562.0 : Bool;   // Bit_00_READY_RUN
   "Carrier_64_G120DStatusWord.1" AT %I3562.1 : Bool;   // Bit_01_READY_ON
   "Carrier_64_G120DStatusWord.2" AT %I3562.2 : Bool;   // Bit_02_ENABLE
   "Carrier_64_G120DStatusWord.3" AT %I3562.3 : Bool;   // Bit_03_FAULT
   "Carrier_64_G120DStatusWord.4" AT %I3562.4 : Bool;   // Bit_04_OFF2
   "Carrier_64_G120DStatusWord.5" AT %I3562.5 : Bool;   // Bit_05_OFF3
   "Carrier_64_G120DStatusWord.6" AT %I3562.6 : Bool;   // Bit_06_LOCK_OUT
   "Carrier_64_G120DStatusWord.7" AT %I3562.7 : Bool;   // Bit_07_WARN
   "Carrier_64_G120DStatusWord.8" AT %I3563.0 : Bool;   // Bit_08_NO_DEVIATION
   "Carrier_64_G120DStatusWord.9" AT %I3563.1 : Bool;   // Bit_09_CONTR_PLC
   "Carrier_64_G120DStatusWord.10" AT %I3563.2 : Bool;   // Bit_10_F_MAX
   "Carrier_64_G120DStatusWord.11" AT %I3563.3 : Bool;   // Bit_11_LIMIT_REACHED
   "Carrier_64_G120DStatusWord.12" AT %I3563.4 : Bool;   // Bit_12_BRAKE_OPEN
   "Carrier_64_G120DStatusWord.13" AT %I3563.5 : Bool;   // Bit_13_NO_OVERTEMP
   "Carrier_64_G120DStatusWord.14" AT %I3563.6 : Bool;   // Bit_14_CW_CCW
   "Carrier_64_G120DStatusWord.15" AT %I3563.7 : Bool;   // Bit_15_OVERL
   "Carrier_64_Slot2_Input" AT %IW3564 : Word;   // SLOT 2 INPUT WORD
   "Carrier_64_CrashDetectSW" AT %I3564.0 : Bool;   // CRASH DETECT SW
   "Carrier_64_SpareSafetyInput(2_1)" AT %I3564.1 : Bool;   // SPARE SAFETY INPUT
   "Carrier_64_SpareSafetyInput(2_2)" AT %I3564.2 : Bool;   // SPARE SAFETY INPUT
   "Carrier_64_SpareSafetyInput(2_3)" AT %I3564.3 : Bool;   // SPARE SAFETY INPUT
   "Carrier_64_SpareSafetyInput(2_4)" AT %I3564.4 : Bool;   // SPARE SAFETY INPUT
   "Carrier_64_SpareSafetyInput(2_5)" AT %I3564.5 : Bool;   // SPARE SAFETY INPUT
   "Carrier_64_SpareSafetyInput(2_6)" AT %I3564.6 : Bool;   // SPARE SAFETY INPUT
   "Carrier_64_SpareSafetyInput(2_7)" AT %I3564.7 : Bool;   // SPARE SAFETY INPUT
   "Carrier_64_Slot3_SafetyOutput" AT %IW3565 : Word;   // SLOT 3 SAFETY OUTPUT WORD
   "Carrier_64_Crash_Detect_OK" AT %I3565.0 : Bool;   // CARRIER CRASH DETECT
   "Carrier_64_SpareSafetyOutput(3_1)" AT %I3565.1 : Bool;   // SPARE SAFETY OUTPUT
   "Carrier_64_SpareSafetyOutput(3_2)" AT %I3565.2 : Bool;   // SPARE SAFETY OUTPUT
   "Carrier_64_SpareSafetyOutput(3_3)" AT %I3565.3 : Bool;   // SPARE SAFETY OUTPUT
   "Carrier_64_SpareSafetyOutput(3_4)" AT %I3565.4 : Bool;   // SPARE SAFETY OUTPUT
   "Carrier_64_SpareSafetyOutput(3_5)" AT %I3565.5 : Bool;   // SPARE SAFETY OUTPUT
   "Carrier_64_SpareSafetyOutput(3_6)" AT %I3565.6 : Bool;   // SPARE SAFETY OUTPUT
   "Carrier_64_SpareSafetyOutput(3_7)" AT %I3565.7 : Bool;   // SPARE SAFETY OUTPUT
   "Carrier_64_Slot4_Input" AT %IW3566 : Word;   // SLOT 4 INPUT WORD
   "Carrier_64_480VPowerOn_MDCB1" AT %I3566.0 : Bool;   // 480 VAC POWER ON MDCB 1
   "Carrier_64_SpareInput(4_1)" AT %I3566.1 : Bool;   // SPARE INPUT
   "Carrier_64_SpareInput(4_2)" AT %I3566.2 : Bool;   // SPARE INPUT
   "Carrier_64_SitopSelectStatus" AT %I3566.3 : Bool;   // SITOP SELECT STATUS
   "Carrier_64_DCsupplyOnPSCB2" AT %I3566.4 : Bool;   // DC SUPPLY ON PSCB 2
   "Carrier_64_SpareInput(4_5)" AT %I3566.5 : Bool;   // SPARE INPUT
   "Carrier_64_SpareInput(4_6)" AT %I3566.6 : Bool;   // SPARE INPUT
   "Carrier_64_SpareInput(4_7)" AT %I3566.7 : Bool;   // SPARE INPUT
   "Carrier_64_PB1_ProdHoldLH" AT %I3567.0 : Bool;   // PB 1 PRODUCTION HOLD LH
   "Carrier_64_PB2_ResetLH" AT %I3567.1 : Bool;   // PB 2 RESET LH
   "Carrier_64_PB3_ProdHoldRH" AT %I3567.2 : Bool;   // PB 3 PRODUCTION HOLD RH
   "Carrier_64_PB4_ResetRH" AT %I3567.3 : Bool;   // PB 4 RESET RH
   "Carrier_64_SpareInput(4_14)" AT %I3567.4 : Bool;   // SPARE INPUT
   "Carrier_64_SpareInput(4_15)" AT %I3567.5 : Bool;   // SPARE INPUT
   "Carrier_64_SpareInput(4_16)" AT %I3567.6 : Bool;   // SPARE INPUT
   "Carrier_64_SpareInput(4_17)" AT %I3567.7 : Bool;   // SPARE INPUT
   "Carrier_64_Slot5_Output" AT %IW3568 : Word;   // SLOT 5 OUTPUT WORD
   "Carrier_64_IRD400_HMI_24VDC_ENABLE" AT %I3568.0 : Bool;   // IRD 400 PANEL HMI 24V DC POWER
   "Carrier_64_FaultLight_LH" AT %I3568.1 : Bool;   // FAULT LIGHT LH
   "Carrier_64_RunLight_LH" AT %I3568.2 : Bool;   // RUN LIGHT LH
   "Carrier_64_FaultLight_RH" AT %I3568.3 : Bool;   // FAULT LIGHT RH
   "Carrier_64_RunLight_RH" AT %I3568.4 : Bool;   // RUN LIGHT RH
   "Carrier_64_SpareOutput(5_5)" AT %I3568.5 : Bool;   // SPARE OUTPUT
   "Carrier_64_SpareOutput(5_6)" AT %I3568.6 : Bool;   // SPARE OUTPUT
   "Carrier_64_SpareOutput(5_7)" AT %I3568.7 : Bool;   // SPARE OUTPUT
   "Carrier_64_ActualSpeed" AT %IW3570 : Word;   // ACTUAL SPEED
   "Carrier_64_CarrierDriveAlarm" AT %IW3572 : Word;   // CARRIER DRIVE ALARM
   "Carrier_64_CarrierDriveWarning" AT %IW3574 : Word;   // CARRIER DRIVE WARNING
   "Carrier_65_Status" AT %IW3600 : Word;   // CARRIER STATUS WORD
   "Carrier_65_Status.0" AT %I3600.0 : Bool;   // HEARTBEAT
   "Carrier_65_Status.1" AT %I3600.1 : Bool;   // MANUAL
   "Carrier_65_Status.2" AT %I3600.2 : Bool;   // IN_AUTO